   "IA Compressor Shutdown Active" : Bool = PLC "10 DI_DATA".E131_SHTDN AT %DB1.DBX0.0, 1 s
   "IDB_ATO2B_1_HIGH LEVEL VALUE (H)" : Real = PLC IDB_ATO2B_1."HIGH LEVEL VALUE (H)" AT %DB731.DBD30, 1 s
   "IDB_ATO2B_1_LOW LEVEL VALUE (L)" : Real = PLC IDB_ATO2B_1."LOW LEVEL VALUE (L)" AT %DB731.DBD26, 1 s
   "IDB_ATO2B_1_VERY HIGH LEVEL VALUE (HH)" : Real = PLC IDB_ATO2B_1."VERY HIGH LEVEL VALUE (HH)" AT %DB731.DBD34, 1 s
   "IDB_ATO2B_1_VERY LOW LEVEL VALUE (LL)" : Real = PLC IDB_ATO2B_1."VERY LOW LEVEL VALUE (LL)" AT %DB731.DBD22, 1 s
   "IDB_E-600_HIGH LEVEL VALUE (H)" : Real = PLC "IDB_E-600"."HIGH LEVEL VALUE (H)" AT %DB600.DBD30, 1 s
   "IDB_E-600_LOW LEVEL VALUE (L)" : Real = PLC "IDB_E-600"."LOW LEVEL VALUE (L)" AT %DB600.DBD26, 1 s
   "IDB_E-600_VERY HIGH LEVEL VALUE (HH)" : Real = PLC "IDB_E-600"."VERY HIGH LEVEL VALUE (HH)" AT %DB600.DBD34, 1 s
   "IDB_E-600_VERY LOW LEVEL VALUE (LL)" : Real = PLC "IDB_E-600"."VERY LOW LEVEL VALUE (LL)" AT %DB600.DBD22, 1 s
   "IDB_E700 Alarms_HIGH LEVEL VALUE (H)" : Real = PLC "IDB_E700 Alarms"."HIGH LEVEL VALUE (H)" AT %DB701.DBD30, 1 s
   "IDB_E700 Alarms_LOW LEVEL VALUE (L)" : Real = PLC "IDB_E700 Alarms"."LOW LEVEL VALUE (L)" AT %DB701.DBD26, 1 s
   "IDB_E700 Alarms_VERY HIGH LEVEL VALUE (HH)" : Real = PLC "IDB_E700 Alarms"."VERY HIGH LEVEL VALUE (HH)" AT %DB701.DBD34, 1 s
   "IDB_E700 Alarms_VERY LOW LEVEL VALUE (LL)" : Real = PLC "IDB_E700 Alarms"."VERY LOW LEVEL VALUE (LL)" AT %DB701.DBD22, 1 s
   "IDB_PIT 102_HIGH LEVEL VALUE (H)" : Real = PLC "IDB_PIT 102"."HIGH LEVEL VALUE (H)" AT %DB722.DBD30, 1 s
   "IDB_PIT 102_LOW LEVEL VALUE (L)" : Real = PLC "IDB_PIT 102"."LOW LEVEL VALUE (L)" AT %DB722.DBD26, 1 s
   "IDB_PIT 102_VERY HIGH LEVEL VALUE (HH)" : Real = PLC "IDB_PIT 102"."VERY HIGH LEVEL VALUE (HH)" AT %DB722.DBD34, 1 s
   "IDB_PIT 102_VERY LOW LEVEL VALUE (LL)" : Real = PLC "IDB_PIT 102"."VERY LOW LEVEL VALUE (LL)" AT %DB722.DBD22, 1 s
   "IDB_PIT 204_HIGH LEVEL VALUE (H)" : Real = PLC "IDB_PIT 204"."HIGH LEVEL VALUE (H)" AT %DB724.DBD30, 1 s
   "IDB_PIT 204_LOW LEVEL VALUE (L)" : Real = PLC "IDB_PIT 204"."LOW LEVEL VALUE (L)" AT %DB724.DBD26, 1 s
   "IDB_PIT 204_VERY HIGH LEVEL VALUE (HH)" : Real = PLC "IDB_PIT 204"."VERY HIGH LEVEL VALUE (HH)" AT %DB724.DBD34, 1 s
   "IDB_PIT 204_VERY LOW LEVEL VALUE (LL)" : Real = PLC "IDB_PIT 204"."VERY LOW LEVEL VALUE (LL)" AT %DB724.DBD22, 1 s
   "IDB_PIT 316_HIGH LEVEL VALUE (H)" : Real = PLC "IDB_PIT 316"."HIGH LEVEL VALUE (H)" AT %DB716.DBD30, 1 s
   "IDB_PIT 316_LOW LEVEL VALUE (L)" : Real = PLC "IDB_PIT 316"."LOW LEVEL VALUE (L)" AT %DB716.DBD26, 1 s
   "IDB_PIT 316_VERY HIGH LEVEL VALUE (HH)" : Real = PLC "IDB_PIT 316"."VERY HIGH LEVEL VALUE (HH)" AT %DB716.DBD34, 1 s
   "IDB_PIT 316_VERY LOW LEVEL VALUE (LL)" : Real = PLC "IDB_PIT 316"."VERY LOW LEVEL VALUE (LL)" AT %DB716.DBD22, 1 s
   "IDB_PIT 359_HIGH LEVEL VALUE (H)" : Real = PLC "IDB_PIT 359"."HIGH LEVEL VALUE (H)" AT %DB759.DBD30, 1 s
   "IDB_PIT 359_LOW LEVEL VALUE (L)" : Real = PLC "IDB_PIT 359"."LOW LEVEL VALUE (L)" AT %DB759.DBD26, 1 s
   "IDB_PIT 359_VERY HIGH LEVEL VALUE (HH)" : Real = PLC "IDB_PIT 359"."VERY HIGH LEVEL VALUE (HH)" AT %DB759.DBD34, 1 s
   "IDB_PIT 359_VERY LOW LEVEL VALUE (LL)" : Real = PLC "IDB_PIT 359"."VERY LOW LEVEL VALUE (LL)" AT %DB759.DBD22, 1 s
   "IDB_PIT 402_HIGH LEVEL VALUE (H)" : Real = PLC "IDB_PIT 402"."HIGH LEVEL VALUE (H)" AT %DB742.DBD30, 1 s
   "IDB_PIT 402_LOW LEVEL VALUE (L)" : Real = PLC "IDB_PIT 402"."LOW LEVEL VALUE (L)" AT %DB742.DBD26, 1 s
   "IDB_PIT 402_VERY HIGH LEVEL VALUE (HH)" : Real = PLC "IDB_PIT 402"."VERY HIGH LEVEL VALUE (HH)" AT %DB742.DBD34, 1 s
   "IDB_PIT 402_VERY LOW LEVEL VALUE (LL)" : Real = PLC "IDB_PIT 402"."VERY LOW LEVEL VALUE (LL)" AT %DB742.DBD22, 1 s
   "IDB_TIT 315_HIGH LEVEL VALUE (H)" : Real = PLC "IDB_TIT 315"."HIGH LEVEL VALUE (H)" AT %DB715.DBD30, 1 s
   "IDB_TIT 315_LOW LEVEL VALUE (L)" : Real = PLC "IDB_TIT 315"."LOW LEVEL VALUE (L)" AT %DB715.DBD26, 1 s
   "IDB_TIT 315_VERY HIGH LEVEL VALUE (HH)" : Real = PLC "IDB_TIT 315"."VERY HIGH LEVEL VALUE (HH)" AT %DB715.DBD34, 1 s
   "IDB_TIT 315_VERY LOW LEVEL VALUE (LL)" : Real = PLC "IDB_TIT 315"."VERY LOW LEVEL VALUE (LL)" AT %DB715.DBD22, 1 s
   "IDB_TIT 319_HIGH LEVEL VALUE (H)" : Real = PLC "IDB_TIT 319"."HIGH LEVEL VALUE (H)" AT %DB719.DBD30, 1 s
   "IDB_TIT 319_LOW LEVEL VALUE (L)" : Real = PLC "IDB_TIT 319"."LOW LEVEL VALUE (L)" AT %DB719.DBD26, 1 s
   "IDB_TIT 319_VERY HIGH LEVEL VALUE (HH)" : Real = PLC "IDB_TIT 319"."VERY HIGH LEVEL VALUE (HH)" AT %DB719.DBD34, 1 s
   "IDB_TIT 319_VERY LOW LEVEL VALUE (LL)" : Real = PLC "IDB_TIT 319"."VERY LOW LEVEL VALUE (LL)" AT %DB719.DBD22, 1 s
   "IDB_TIT 360_HIGH LEVEL VALUE (H)" : Real = PLC "IDB_TIT 360"."HIGH LEVEL VALUE (H)" AT %DB760.DBD30, 1 s
   "IDB_TIT 360_LOW LEVEL VALUE (L)" : Real = PLC "IDB_TIT 360"."LOW LEVEL VALUE (L)" AT %DB760.DBD26, 1 s
   "IDB_TIT 360_VERY HIGH LEVEL VALUE (HH)" : Real = PLC "IDB_TIT 360"."VERY HIGH LEVEL VALUE (HH)" AT %DB760.DBD34, 1 s
   "IDB_TIT 360_VERY LOW LEVEL VALUE (LL)" : Real = PLC "IDB_TIT 360"."VERY LOW LEVEL VALUE (LL)" AT %DB760.DBD22, 1 s
   "IDB_TIT 401_HIGH LEVEL VALUE (H)" : Real = PLC "IDB_TIT 401"."HIGH LEVEL VALUE (H)" AT %DB741.DBD30, 1 s
   "IDB_TIT 401_LOW LEVEL VALUE (L)" : Real = PLC "IDB_TIT 401"."LOW LEVEL VALUE (L)" AT %DB741.DBD26, 1 s
   "IDB_TIT 401_VERY HIGH LEVEL VALUE (HH)" : Real = PLC "IDB_TIT 401"."VERY HIGH LEVEL VALUE (HH)" AT %DB741.DBD34, 1 s
   "IDB_TIT 401_VERY LOW LEVEL VALUE (LL)" : Real = PLC "IDB_TIT 401"."VERY LOW LEVEL VALUE (LL)" AT %DB741.DBD22, 1 s
   "IG Press SP (R)" : Real = PLC "19_AUTO_CMNDS_Data".PIT402_Target AT %DB1.DBD0, 1 s
   "IG Shell Temp Hi Switch" : Bool = PLC "10 DI_DATA".TS006 AT %DB1.DBX0.0, 1 s
   "IG Soot Content Scaled" : Real = PLC "12_AI_Data".E700SootContentIn AT %DB1.DBX0.0, 1 s
   "IG Temp Hi Hi Switch" : Bool = PLC "10 DI_DATA".TS403_FAULT AT %DB1.DBX0.0, 1 s
   "IG Temperature High (TS403)" : Bool = PLC "10 DI_DATA".TS403_FAULT AT %DB1.DBX0.0, 1 s
   "IGG Automated" : Bool = PLC "80_From_HMI".Request_Auto AT %DB1.DBX0.0, 1 s
   "IGG E-Stop Healthy" : Bool = PLC "10_DI_Data".IGG_ESTOP_OK AT %DB1.DBX0.0, 1 s
   "IGG Inlet Fuel Pressure (PIT204) Scaled" : Real = PLC "12_AI_Data".PIT204In_SCALED AT %DB1.DBX0.0, 1 s
   "IGG Inlet Fuel Temp (TIT202) Scaled" : Real = PLC "12_AI_Data".TIT202In_SCALED AT %DB1.DBX0.0, 1 s
   "IGG Main Atom Air Presure (PIT113) Scaled" : Real = PLC "12_AI_Data".PIT113In_SCALED AT %DB1.DBX0.0, 1 s
   "IGG Main Fuel Pressure (PIT205) Scaled" : Real = PLC "12_AI_Data".PIT205In_SCALED AT %DB1.DBX0.0, 1 s
   "IGG Manual" : Bool = PLC "80_From_HMI".Request_Manual AT %DB1.DBX0.0, 1 s
   "IGG Running" : Bool = PLC "14_DQ_Data".24PF1 AT %DB1.DBX0.0, 1 s
   "IGG Shell High Temp (TS006)" : Bool = PLC "10 DI_DATA".TS006 AT %DB1.DBX0.0, 1 s
   "IGG Shutdown Alarm Active" : Bool = PLC "14_DQ_Data".24K3 AT %DB1.DBX0.0, 1 s
   "IGG Shutting Down animation" : Bool = PLC "14_DQ_Data".24K3 AT %DB1.DBX0.0, 1 s
   "IGG Start Warning" : Bool = PLC "Sequence Times_DB"."Warn to IGG Start" AT %DB1.DBW0, 1 s
   "IGG Vent Power Healthy" : Bool = PLC "10_DI_Data".IGG_VNT_PWR_OK AT %DB1.DBX0.0, 1 s
   "IGG Warning Alarm Active" : Bool = PLC "14_DQ_Data".24K4 AT %DB1.DBX0.0, 1 s
   "IGG_Step_Time_001" : Time = PLC "86_Times".STEP_MAX_TIME_STP_001 AT %DB1.DBW0, 1 s
   "IGG_Step_Time_005" : Time = PLC "86_Times".STEP_MAX_TIME_STP_005 AT %DB1.DBW0, 1 s
   "IGG_Step_Time_010" : Time = PLC "86_Times".STEP_MAX_TIME_STP_010 AT %DB1.DBW0, 1 s
   "IGG_Step_Time_020" : Time = PLC "86_Times".STEP_MAX_TIME_STP_020 AT %DB1.DBW0, 1 s
   "IGG_Step_Time_030" : Time = PLC "86_Times".STEP_MAX_TIME_STP_030 AT %DB1.DBW0, 1 s
   "IGG_Step_Time_040" : Time = PLC "86_Times".STEP_MAX_TIME_STP_040 AT %DB1.DBW0, 1 s
   "IGG_Step_Time_050" : Time = PLC "86_Times".STEP_MAX_TIME_STP_050 AT %DB1.DBW0, 1 s
   "IGG_Step_Time_060" : Time = PLC "86_Times".STEP_MAX_TIME_STP_060 AT %DB1.DBW0, 1 s
   "IGG_Step_Time_070" : Time = PLC "86_Times".STEP_MAX_TIME_STP_070 AT %DB1.DBW0, 1 s
   "IGG_Step_Time_080" : Time = PLC "86_Times".STEP_MAX_TIME_STP_080 AT %DB1.DBW0, 1 s
   "IGG_Step_Time_090" : Time = PLC "86_Times".STEP_MAX_TIME_STP_090 AT %DB1.DBW0, 1 s
   "IGG_Step_Time_100" : Time = PLC "86_Times".STEP_MAX_TIME_STP_100 AT %DB1.DBW0, 1 s
   "IGG_Step_Time_110" : Time = PLC "86_Times".STEP_MAX_TIME_STP_110 AT %DB1.DBW0, 1 s
   "IGG_Step_Time_120" : Time = PLC "86_Times".STEP_MAX_TIME_STP_120 AT %DB1.DBW0, 1 s
   "IGG_Step_Time_130" : Time = PLC "86_Times".STEP_MAX_TIME_STP_130 AT %DB1.DBW0, 1 s
   "IGG_Step_Time_140" : Time = PLC "86_Times".STEP_MAX_TIME_STP_140 AT %DB1.DBW0, 1 s
   "IGG_Step_Time_150" : Time = PLC "86_Times".STEP_MAX_TIME_STP_150 AT %DB1.DBW0, 1 s
   "IGG_Step_Time_160" : Time = PLC "86_Times".STEP_MAX_TIME_STP_160 AT %DB1.DBW0, 1 s
   "IGG_Step_Time_170" : Time = PLC "86_Times".STEP_MAX_TIME_STP_170 AT %DB1.DBW0, 1 s
   "IGG_Step_Time_180" : Time = PLC "86_Times".STEP_MAX_TIME_STP_180 AT %DB1.DBW0, 1 s
   "IGG_Step_Time_190" : Time = PLC "86_Times".STEP_MAX_TIME_STP_190 AT %DB1.DBW0, 1 s
   "IGG_Step_Time_200" : Time = PLC "86_Times".STEP_MAX_TIME_STP_200 AT %DB1.DBW0, 1 s
   "IGG_Step_Time_210" : Time = PLC "86_Times".STEP_MAX_TIME_STP_210 AT %DB1.DBW0, 1 s
   "IGG_Step_Time_220" : Time = PLC "86_Times".STEP_MAX_TIME_STP_220 AT %DB1.DBW0, 1 s
   "IGG_Step_Time_230" : Time = PLC "86_Times".STEP_MAX_TIME_STP_230 AT %DB1.DBW0, 1 s
   "IGG_Step_Time_240" : Time = PLC "86_Times".STEP_MAX_TIME_STP_240 AT %DB1.DBW0, 1 s
   "IGG_Step_Time_250" : Time = PLC "86_Times".STEP_MAX_TIME_STP_250 AT %DB1.DBW0, 1 s
   "IGG_Step_Time_260" : Time = PLC "86_Times".STEP_MAX_TIME_STP_260 AT %DB1.DBW0, 1 s
   "IGG_Step_Time_270" : Time = PLC "86_Times".STEP_MAX_TIME_STP_270 AT %DB1.DBW0, 1 s
   "IGG_Step_Time_280" : Time = PLC "86_Times".STEP_MAX_TIME_STP_280 AT %DB1.DBW0, 1 s
   "IGG_Step_Time_290" : Time = PLC "86_Times".STEP_MAX_TIME_STP_290 AT %DB1.DBW0, 1 s
   "IGG_Step_Time_300" : Time = PLC "86_Times".STEP_MAX_TIME_STP_300 AT %DB1.DBW0, 1 s
   "IGG_Step_Time_310" : Time = PLC "86_Times".STEP_MAX_TIME_STP_310 AT %DB1.DBW0, 1 s
   "IGG_Step_Time_320" : Time = PLC "86_Times".STEP_MAX_TIME_STP_320 AT %DB1.DBW0, 1 s
   "IGG_Step_Time_330" : Time = PLC "86_Times".STEP_MAX_TIME_STP_330 AT %DB1.DBW0, 1 s
   "IGG_Step_Time_340" : Time = PLC "86_Times".STEP_MAX_TIME_STP_340 AT %DB1.DBW0, 1 s
   "IGG_Step_Time_350" : Time = PLC "86_Times".STEP_MAX_TIME_STP_350 AT %DB1.DBW0, 1 s
   "IGG_Step_Time_360" : Time = PLC "86_Times".STEP_MAX_TIME_STP_360 AT %DB1.DBW0, 1 s
   "IGG_Step_Time_370" : Time = PLC "86_Times".STEP_MAX_TIME_STP_370 AT %DB1.DBW0, 1 s
   "IGG_Step_Time_380" : Time = PLC "86_Times".STEP_MAX_TIME_STP_380 AT %DB1.DBW0, 1 s
   "IGG_Step_Time_390" : Time = PLC "86_Times".STEP_MAX_TIME_STP_390 AT %DB1.DBW0, 1 s
   "IGG_Step_Time_400" : Time = PLC "86_Times".STEP_MAX_TIME_STP_400 AT %DB1.DBW0, 1 s
   "IGG_Step_Time_410" : Time = PLC "86_Times".STEP_MAX_TIME_STP_410 AT %DB1.DBW0, 1 s
   "IGG_Step_Time_420" : Time = PLC "86_Times".STEP_MAX_TIME_STP_420 AT %DB1.DBW0, 1 s
   "IGG_Step_Time_430" : Time = PLC "86_Times".STEP_MAX_TIME_STP_430 AT %DB1.DBW0, 1 s
   "IGG_Step_Time_440" : Time = PLC "86_Times".STEP_MAX_TIME_STP_440 AT %DB1.DBW0, 1 s
   "IGG_Step_Time_450" : Time = PLC "86_Times".STEP_MAX_TIME_STP_450 AT %DB1.DBW0, 1 s
   "IGG_Step_Time_460" : Time = PLC "86_Times".STEP_MAX_TIME_STP_460 AT %DB1.DBW0, 1 s
   "IGG_Step_Time_470" : Time = PLC "86_Times".STEP_MAX_TIME_STP_470 AT %DB1.DBW0, 1 s
   "IGG_Step_Time_480" : Time = PLC "86_Times".STEP_MAX_TIME_STP_480 AT %DB1.DBW0, 1 s
   "IGG_Step_Time_490" : Time = PLC "86_Times".STEP_MAX_TIME_STP_490 AT %DB1.DBW0, 1 s
   "IGG_Step_Time_500" : Time = PLC "86_Times".STEP_MAX_TIME_STP_500 AT %DB1.DBW0, 1 s
   "IGG_Times_Burner Control Start Command Delay" : Time = PLC "86_Times".PRE_BC_STRT_CMND_DLY AT %DB1.DBD0, 1 s
   "IGG_Times_CV203 Close Command" : Time = PLC "86_Times".PRE_CV203_CLS_CMND_DLY AT %DB1.DBD0, 1 s
   "IGG_Times_CV311 Max" : Time = PLC "86_Times".CV311_MAX_TRVL_TIME AT %DB1.DBD0, 1 s
   "IGG_Times_CV312 Max" : Time = PLC "86_Times".CV312_MAX_TRVL_TIME AT %DB1.DBD0, 1 s
   "IGG_Times_CV321 Max" : Time = PLC "86_Times".CV321_MAX_TRVL_TIME AT %DB1.DBD0, 1 s
   "IGG_Times_CV322 Max" : Time = PLC "86_Times".CV322_MAX_TRVL_TIME AT %DB1.DBD0, 1 s
   "IGG_Times_CV401 Max" : Time = PLC "86_Times".CV401_MAX_TRVL_TIME AT %DB1.DBD0, 1 s
   "IGG_Times_CV431 Max" : Time = PLC "86_Times".CV431_MAX_TRVL_TIME AT %DB1.DBD0, 1 s
   "IGG_Times_CV432 Max" : Time = PLC "86_Times".CV432_MAX_TRVL_TIME AT %DB1.DBD0, 1 s
   "IGG_Times_Post CV311 Close" : Time = PLC "86_Times".POST_CV311_CLS_DLY AT %DB1.DBD0, 1 s
   "IGG_Times_Post CV321 Open" : Time = PLC "86_Times".POST_CV321_OPN_DLY AT %DB1.DBD0, 1 s
   "IGG_Times_Post P301 Stop" : Time = PLC "86_Times".POST_P301_STOP_DLY AT %DB1.DBD0, 1 s
   "Igniter Control" : Bool = PLC "14_DQ_Data".X001ControlOut AT %DB1.DBX0.0, 1 s
   "Ignitor Power Healthy" : Bool = PLC "10 DI_DATA".X001_PWR_OK AT %DB1.DBX0.0, 1 s
   "Inert Gas Pressure (PIT402) Scaled" : Real = PLC "12_AI_Data".PIT402_SCALED AT %DB1.DBX0.0, 1 s
   "Inert Gas Temp Scaled" : Real = PLC "12_AI_Data".TIT401_SCALED AT %DB1.DBX0.0, 1 s
   "Inlet CSW Pressured PIT359 Scaled" : Real = PLC "12_AI_Data".PIT359_SCALED AT %DB1.DBX0.0, 1 s
   "Inlet CSW Temp Scaled" : Real = PLC "12_AI_Data".TIT319_SCALED AT %DB1.DBX0.0, 1 s
   "Inlet IA Pressure PIT112 Scaled" : Real = PLC "12_AI_Data".PIT112In_SCALED AT %DB1.DBX0.0, 1 s
   "Jacket Cooling Water Flow Switch" : Bool = PLC "10 DI_DATA".FS317 AT %DB1.DBX0.0, 1 s
   "LIT304_ALM_ANALOG_DB71_HIGH LEVEL VALUE (H)" : Real = PLC LIT304_ALM_ANALOG_DB71."HIGH LEVEL VALUE (H)" AT %DB71.DBD30, 1 s
   "LIT304_ALM_ANALOG_DB71_LOW LEVEL VALUE (L)" : Real = PLC LIT304_ALM_ANALOG_DB71."LOW LEVEL VALUE (L)" AT %DB71.DBD26, 1 s
   "LIT304_ALM_ANALOG_DB71_VERY HIGH LEVEL VALUE (HH)" : Real = PLC LIT304_ALM_ANALOG_DB71."VERY HIGH LEVEL VALUE (HH)" AT %DB71.DBD34, 1 s
   "LIT304_ALM_ANALOG_DB71_VERY LOW LEVEL VALUE (LL)" : Real = PLC LIT304_ALM_ANALOG_DB71."VERY LOW LEVEL VALUE (LL)" AT %DB71.DBD22, 1 s
   "Logging SD Card Overflow" : Bool AT %DB1.DBX0.0
      on ChangeValue: "SD_Card_Overflow"()
   "Main Atom Air Flow  OK" : Bool = PLC "10 DI_DATA".FS115 AT %DB1.DBX0.0, 1 s
   "Main Atom Air Flow Switch" : Bool = PLC "10 DI_DATA".FS115 AT %DB1.DBW0, 1 s
   "Main Atom Air Reg Valve Position" : Real = PLC "16_AQ_Data".CV111_CNTRL AT %DB1.DBD0, 1 s
   "Main B Atom Air Valve Control" : Bool = PLC "14_DQ_Data".200CV114ControlOut AT %DB1.DBX0.0, 1 s
   "Main B Fuel Valve 1 Control" : Bool = PLC "14_DQ_Data".200CV206ControlOut AT %DB1.DBX0.0, 1 s
   "Main B Fuel Valve 2 Control" : Bool = PLC "14_DQ_Data".200CV207ControlOut AT %DB1.DBX0.0, 1 s
   "Main Fuel Reg Valve Control" : Real = PLC "16_AQ_Data".CV203_CNTRL AT %DB1.DBD0, 1 s
   "Main Fuel Reg Valve Position" : Real = PLC "16_AQ_Data".CV203_CNTRL, 1 s
   "Maintained 24V Power" : Bool = PLC "10_DI_Data".MAINTD_24VDC_PWR_OK AT %DB1.DBX0.0, 1 s
   "MAN_AQ100_DEC_CAB_Speed" : Bool = PLC "80_From_HMI".MAN_AQ_DEC_100 AT %DB1.DBX0.0, 1 s
   "MAN_AQ100_DEC_Main_Fuel_Reg" : Bool = PLC "80_From_HMI".MAN_AQ_DEC_100 AT %DB1.DBX0.0, 1 s
   "MAN_AQ100_INC_CAB_Speed" : Bool = PLC "80_From_HMI".MAN_AQ_INC_100 AT %DB1.DBX0.0, 1 s
   "MAN_AQ100_INC_Main_Fuel_Reg" : Bool = PLC "80_From_HMI".MAN_AQ_INC_100 AT %DB1.DBX0.0, 1 s
   "MAN_AQ102_DEC_Main_Atom_Air" : Bool = PLC "80_From_HMI".MAN_AQ_DEC_102 AT %DB1.DBX0.0, 1 s
   "MAN_AQ102_DEC_SPARE" : Bool = PLC "80_From_HMI".MAN_AQ_DEC_102 AT %DB1.DBX0.0, 1 s
   "MAN_AQ102_INC_Main_Atom_Air" : Bool = PLC "80_From_HMI".MAN_AQ_INC_102 AT %DB1.DBX0.0, 1 s
   "MAN_AQ102_INC_SPARE" : Bool = PLC "80_From_HMI".MAN_AQ_INC_102 AT %DB1.DBX0.0, 1 s
   "MAN_AQ104_DEC_SPARE" : Bool = PLC "80_From_HMI".MAN_AQ_DEC_104 AT %DB1.DBX0.0, 1 s
   "MAN_AQ104_INC_SPARE" : Bool = PLC "80_From_HMI".MAN_AQ_INC_104 AT %DB1.DBX0.0, 1 s
   "MAN_AQ96_DEC_SPARE" : Bool = PLC "80_From_HMI".MAN_AQ_DEC_96 AT %DB1.DBX0.0, 1 s
   "MAN_AQ96_INC_SPARE" : Bool = PLC "80_From_HMI".MAN_AQ_INC_96 AT %DB1.DBX0.0, 1 s
   "MAN_AQ98_DEC_SPARE" : Bool = PLC "80_From_HMI".MAN_AQ_DEC_98 AT %DB1.DBX0.0, 1 s
   "MAN_AQ98_DEC_Vent_Valve_Pos" : Bool = PLC "80_From_HMI".MAN_AQ_DEC_98 AT %DB1.DBX0.0, 1 s
   "MAN_AQ98_INC_SPARE" : Bool = PLC "80_From_HMI".MAN_AQ_INC_98 AT %DB1.DBX0.0, 1 s
   "MAN_AQ98_INC_Vent_Valve_Pos" : Bool = PLC "80_From_HMI".MAN_AQ_INC_98 AT %DB1.DBX0.0, 1 s
   "MAN_Q0.0_FP1" : Bool = PLC "80_From_HMI".MAN_DQ_0_0 AT %DB1.DBX0.0, 1 s
   "MAN_Q0.0_Test_Press" : Bool = PLC "80_From_HMI".MAN_DQ_0_0 AT %DB1.DBX0.0, 1 s
   "MAN_Q0.1_FP2" : Bool = PLC "80_From_HMI".MAN_DQ_0_1 AT %DB1.DBX0.0, 1 s
   "MAN_Q0.1_Pilot_IGN" : Bool = PLC "80_From_HMI".MAN_DQ_0_1 AT %DB1.DBX0.0, 1 s
   "MAN_Q0.2_CAB" : Bool = PLC "80_From_HMI".MAN_DQ_0_2 AT %DB1.DBX0.0, 1 s
   "MAN_Q0.2_PilotFuel1" : Bool = PLC "80_From_HMI".MAN_DQ_0_2 AT %DB1.DBX0.0, 1 s
   "MAN_Q0.3_CSW_Inlet" : Bool = PLC "80_From_HMI".MAN_DQ_0_3 AT %DB1.DBX0.0, 1 s
   "MAN_Q0.3_PilotFuel2" : Bool = PLC "80_From_HMI".MAN_DQ_0_3 AT %DB1.DBX0.0, 1 s
   "MAN_Q0.4_CSW_Drain" : Bool = PLC "80_From_HMI".MAN_DQ_0_4 AT %DB1.DBX0.0, 1 s
   "MAN_Q0.4_MainAtom" : Bool = PLC "80_From_HMI".MAN_DQ_0_4 AT %DB1.DBX0.0, 1 s
   "MAN_Q0.5_IGSupply" : Bool = PLC "80_From_HMI".MAN_DQ_0_5 AT %DB1.DBX0.0, 1 s
   "MAN_Q0.5_MainFuel1" : Bool = PLC "80_From_HMI".MAN_DQ_0_5 AT %DB1.DBX0.0, 1 s
   "MAN_Q0.6_CB/BWTS" : Bool = PLC "80_From_HMI".MAN_DQ_0_6 AT %DB1.DBX0.0, 1 s
   "MAN_Q0.6_MainFuel2" : Bool = PLC "80_From_HMI".MAN_DQ_0_6 AT %DB1.DBX0.0, 1 s
   "MAN_Q0.7_IAComp" : Bool = PLC "80_From_HMI".MAN_DQ_0_7 AT %DB1.DBX0.0, 1 s
   "MAN_Q0.7_Spare" : Bool = PLC "80_From_HMI".MAN_DQ_0_7 AT %DB1.DBX0.0, 1 s
   "MAN_Q1.0_CSWPump" : Bool = PLC "80_From_HMI".MAN_DQ_1_0 AT %DB1.DBX0.0, 1 s
   "MAN_Q1.0_Spare" : Bool = PLC "80_From_HMI".MAN_DQ_1_0 AT %DB1.DBX0.0, 1 s
   "MAN_Q1.1_Atmos" : Bool = PLC "80_From_HMI".MAN_DQ_1_1 AT %DB1.DBX0.0, 1 s
   "MAN_Q1.1_IGN" : Bool = PLC "80_From_HMI".MAN_DQ_1_1 AT %DB1.DBX0.0, 1 s
   "MAN_Q1.2_IGG_SD" : Bool = PLC "80_From_HMI".MAN_DQ_1_2 AT %DB1.DBX0.0, 1 s
   "MAN_Q1.2_Spare" : Bool = PLC "80_From_HMI".MAN_DQ_1_2 AT %DB1.DBX0.0, 1 s
   "MAN_Q1.3_IGG_WRN" : Bool = PLC "80_From_HMI".MAN_DQ_1_3 AT %DB1.DBX0.0, 1 s
   "MAN_Q1.3_Spare" : Bool = PLC "80_From_HMI".MAN_DQ_1_3 AT %DB1.DBX0.0, 1 s
   "MAN_Q1.4_IGG_RNG" : Bool = PLC "80_From_HMI".MAN_DQ_1_4 AT %DB1.DBX0.0, 1 s
   "MAN_Q1.4_Spare" : Bool = PLC "80_From_HMI".MAN_DQ_1_4 AT %DB1.DBX0.0, 1 s
   "MAN_Q1.5_SD" : Bool = PLC "80_From_HMI".MAN_DQ_1_5 AT %DB1.DBX0.0, 1 s
   "MAN_Q1.5_Spare" : Bool = PLC "80_From_HMI".MAN_DQ_1_5 AT %DB1.DBX0.0, 1 s
   "MAN_Q1.6_Spare" : Bool = PLC "80_From_HMI".MAN_DQ_1_6 AT %DB1.DBX0.0, 1 s
   "MAN_Q1.6_WRN" : Bool = PLC "80_From_HMI".MAN_DQ_1_6 AT %DB1.DBX0.0, 1 s
   "MAN_Q1.7_BUZ" : Bool = PLC "80_From_HMI".MAN_DQ_1_7 AT %DB1.DBX0.0, 1 s
   "MAN_Q1.7_CSW_Pump" : Bool = PLC "80_From_HMI".MAN_DQ_1_7 AT %DB1.DBX0.0, 1 s
   "MCC Vent Power Healthy" : Bool = PLC "10_DI_Data".MCC_VNT_PWR_OK AT %DB1.DBX0.0, 1 s
   "Not BWT mode Warning" : Bool = PLC "2068_Sys_Status_Data"."Not BWT mode Warning" AT %DB1.DBD0, 1 s
   "Nozzle Cooling Water Flow Switch" : Bool = PLC "10 DI_DATA".FS320 AT %DB1.DBX0.0, 1 s
   "O2 Analyser Content Scaled" : Real = PLC "12_AI_Data".E600O2ContentIn AT %DB1.DBX0.0, 100 ms
   "O2 Analyser Hi Hi" : Bool = PLC "10 DI_DATA".E600_HIHI AT %DB1.DBX0.0, 1 s
   "O2 Analyser Lo Lo" : Bool = PLC "10 DI_DATA".E600_LOLO AT %DB1.DBX0.0, 1 s
   "O2 Ramp Control_QLMN_HLM" : Bool = PLC "O2 Ramp Control".QLMN_HLM, 1 s
   "O2 Ramp Control_QLMN_LLM" : Bool = PLC "O2 Ramp Control".QLMN_LLM, 1 s
   "O2 System Fail" : Bool = PLC "10 DI_DATA".E600_NOK AT %DB1.DBX0.0, 1 s
   "O2 System Power Healthy" : Bool = PLC "10 DI_DATA".E600_PWR_OK AT %DB1.DBX0.0, 1 s
   "Operation hours E139_IDB_Hours Functioning" : Int = PLC "Operation hours E139_IDB"."Hours Functioning", 1 s
   "Outlet CSW Pressure PIT316 Scaled" : Real = PLC "12_AI_Data".PIT316_SCALED AT %DB1.DBX0.0, 1 s
   "Outlet CSW Temp Scaled" : Real = PLC "12_AI_Data".TIT360_SCALED AT %DB1.DBX0.0, 1 s
   "P301 Present" : Bool = PLC "80_From_HMI".P301_PRSNT AT %DB1.DBX0.0, 1 s
   "P305_Functioning Hours_IDB_Hours Functioning Out" : Int = PLC "P305_Functioning Hours_IDB"."Hours Functioning Out", 1 s
   "PGC_COMMISSION_MODE_DB_Active" : Bool = PLC PGC_COMMISSION_MODE_DB.Active, 1 s
   "PGC_COMMISSION_MODE_DB_Button Control" : Int = PLC PGC_COMMISSION_MODE_DB."Button Control", 1 s
   "PGC_COMMISSION_MODE_DB_Drive Popup" : Bool = PLC PGC_COMMISSION_MODE_DB."Drive Popup", 500 ms
   "PGC_COMMISSION_MODE_DB_Setpoint" : Real = PLC PGC_COMMISSION_MODE_DB.Setpoint, 1 s
   "Pilot Air Flow  OK" : Bool = PLC "10 DI_DATA".FS123 AT %DB1.DBX0.0, 1 s
   "Pilot B Fuel Valve 1 Control" : Bool = PLC "14_DQ_Data".200CV215ControlOut AT %DB1.DBX0.0, 1 s
   "Pilot B Fuel Valve 2 Control" : Bool = PLC "14_DQ_Data".200CV216ControlOut AT %DB1.DBX0.0, 1 s
   "Pilot B Ignition Air Valve Control" : Bool = PLC "14_DQ_Data".200CV124ControlOut AT %DB1.DBX0.0, 1 s
   "Pilot Flame" : Bool = PLC "102_Pilot_Burner_DB".FLM_DET AT %DB1.DBX0.0, 100 ms
   "PilotPurgeOK" : Bool = PLC "104_Pilot_Purge_DB".DN_OK AT %DB1.DBX0.0, 1 s
   "PIT348_ALM_ANALOG_DB73_HIGH LEVEL VALUE (H)" : Real = PLC PIT348_ALM_ANALOG_DB73."HIGH LEVEL VALUE (H)" AT %DB73.DBD30, 1 s
   "PIT348_ALM_ANALOG_DB73_LOW LEVEL VALUE (L)" : Real = PLC PIT348_ALM_ANALOG_DB73."LOW LEVEL VALUE (L)" AT %DB73.DBD26, 1 s
   "PIT348_ALM_ANALOG_DB73_VERY HIGH LEVEL VALUE (HH)" : Real = PLC PIT348_ALM_ANALOG_DB73."VERY HIGH LEVEL VALUE (HH)" AT %DB73.DBD34, 1 s
   "PIT348_ALM_ANALOG_DB73_VERY LOW LEVEL VALUE (LL)" : Real = PLC PIT348_ALM_ANALOG_DB73."VERY LOW LEVEL VALUE (LL)" AT %DB73.DBD22, 1 s
   "PIT353_ALM_ANALOG_DB72_HIGH LEVEL VALUE (H)" : Real = PLC PIT353_ALM_ANALOG_DB72."HIGH LEVEL VALUE (H)" AT %DB72.DBD30, 1 s
   "PIT353_ALM_ANALOG_DB72_LOW LEVEL VALUE (L)" : Real = PLC PIT353_ALM_ANALOG_DB72."LOW LEVEL VALUE (L)" AT %DB72.DBD26, 1 s
   "PIT353_ALM_ANALOG_DB72_VERY HIGH LEVEL VALUE (HH)" : Real = PLC PIT353_ALM_ANALOG_DB72."VERY HIGH LEVEL VALUE (HH)" AT %DB72.DBD34, 1 s
   "PIT353_ALM_ANALOG_DB72_VERY LOW LEVEL VALUE (LL)" : Real = PLC PIT353_ALM_ANALOG_DB72."VERY LOW LEVEL VALUE (LL)" AT %DB72.DBD22, 1 s
   "PIT358_ALM_ANALOG_DB78_HIGH LEVEL VALUE (H)" : Real = PLC PIT358_ALM_ANALOG_DB78."HIGH LEVEL VALUE (H)" AT %DB78.DBD30, 1 s
   "PIT358_ALM_ANALOG_DB78_LOW LEVEL VALUE (L)" : Real = PLC PIT358_ALM_ANALOG_DB78."LOW LEVEL VALUE (L)" AT %DB78.DBD26, 1 s
   "PIT358_ALM_ANALOG_DB78_VERY HIGH LEVEL VALUE (HH)" : Real = PLC PIT358_ALM_ANALOG_DB78."VERY HIGH LEVEL VALUE (HH)" AT %DB78.DBD34, 1 s
   "PIT358_ALM_ANALOG_DB78_VERY LOW LEVEL VALUE (LL)" : Real = PLC PIT358_ALM_ANALOG_DB78."VERY LOW LEVEL VALUE (LL)" AT %DB78.DBD22, 1 s
   "PIT424_RIO1_ALM_ANALOG_DB_HIGH LEVEL VALUE (H)" : Real = PLC PIT424_RIO1_ALM_ANALOG_DB."HIGH LEVEL VALUE (H)" AT %DB2219.DBD30, 1 s
   "PIT424_RIO1_ALM_ANALOG_DB_LOW LEVEL VALUE (L)" : Real = PLC PIT424_RIO1_ALM_ANALOG_DB."LOW LEVEL VALUE (L)" AT %DB2219.DBD26, 1 s
   "PIT424_RIO1_ALM_ANALOG_DB_VERY HIGH LEVEL VALUE (HH)" : Real = PLC PIT424_RIO1_ALM_ANALOG_DB."VERY HIGH LEVEL VALUE (HH)" AT %DB2219.DBD34, 1 s
   "PIT424_RIO1_ALM_ANALOG_DB_VERY LOW LEVEL VALUE (LL)" : Real = PLC PIT424_RIO1_ALM_ANALOG_DB."VERY LOW LEVEL VALUE (LL)" AT %DB2219.DBD22, 1 s
   "PIT424_RIO3_ALM_ANALOG_DB_HIGH LEVEL VALUE (H)" : Real = PLC PIT424_RIO3_ALM_ANALOG_DB."HIGH LEVEL VALUE (H)" AT %DB2220.DBD30, 1 s
   "PIT424_RIO3_ALM_ANALOG_DB_LOW LEVEL VALUE (L)" : Real = PLC PIT424_RIO3_ALM_ANALOG_DB."LOW LEVEL VALUE (L)" AT %DB2220.DBD26, 1 s
   "PIT424_RIO3_ALM_ANALOG_DB_VERY HIGH LEVEL VALUE (HH)" : Real = PLC PIT424_RIO3_ALM_ANALOG_DB."VERY HIGH LEVEL VALUE (HH)" AT %DB2220.DBD34, 1 s
   "PIT424_RIO3_ALM_ANALOG_DB_VERY LOW LEVEL VALUE (LL)" : Real = PLC PIT424_RIO3_ALM_ANALOG_DB."VERY LOW LEVEL VALUE (LL)" AT %DB2220.DBD22, 1 s
   "PIT424_RIO4_ALM_ANALOG_DB_HIGH LEVEL VALUE (H)" : Real = PLC PIT424_RIO4_ALM_ANALOG_DB."HIGH LEVEL VALUE (H)" AT %DB2221.DBD30, 1 s
   "PIT424_RIO4_ALM_ANALOG_DB_LOW LEVEL VALUE (L)" : Real = PLC PIT424_RIO4_ALM_ANALOG_DB."LOW LEVEL VALUE (L)" AT %DB2221.DBD26, 1 s
   "PIT424_RIO4_ALM_ANALOG_DB_VERY HIGH LEVEL VALUE (HH)" : Real = PLC PIT424_RIO4_ALM_ANALOG_DB."VERY HIGH LEVEL VALUE (HH)" AT %DB2221.DBD34, 1 s
   "PIT424_RIO4_ALM_ANALOG_DB_VERY LOW LEVEL VALUE (LL)" : Real = PLC PIT424_RIO4_ALM_ANALOG_DB."VERY LOW LEVEL VALUE (LL)" AT %DB2221.DBD22, 1 s
   "PIT424_RIO5_ALM_ANALOG_DB_HIGH LEVEL VALUE (H)" : Real = PLC PIT424_RIO5_ALM_ANALOG_DB."HIGH LEVEL VALUE (H)" AT %DB2222.DBD30, 1 s
   "PIT424_RIO5_ALM_ANALOG_DB_LOW LEVEL VALUE (L)" : Real = PLC PIT424_RIO5_ALM_ANALOG_DB."LOW LEVEL VALUE (L)" AT %DB2222.DBD26, 1 s
   "PIT424_RIO5_ALM_ANALOG_DB_VERY HIGH LEVEL VALUE (HH)" : Real = PLC PIT424_RIO5_ALM_ANALOG_DB."VERY HIGH LEVEL VALUE (HH)" AT %DB2222.DBD34, 1 s
   "PIT424_RIO5_ALM_ANALOG_DB_VERY LOW LEVEL VALUE (LL)" : Real = PLC PIT424_RIO5_ALM_ANALOG_DB."VERY LOW LEVEL VALUE (LL)" AT %DB2222.DBD22, 1 s
   "PIT424_RIO6_ALM_ANALOG_DB_HIGH LEVEL VALUE (H)" : Real = PLC PIT424_RIO6_ALM_ANALOG_DB."HIGH LEVEL VALUE (H)" AT %DB2223.DBD30, 1 s
   "PIT424_RIO6_ALM_ANALOG_DB_LOW LEVEL VALUE (L)" : Real = PLC PIT424_RIO6_ALM_ANALOG_DB."LOW LEVEL VALUE (L)" AT %DB2223.DBD26, 1 s
   "PIT424_RIO6_ALM_ANALOG_DB_VERY HIGH LEVEL VALUE (HH)" : Real = PLC PIT424_RIO6_ALM_ANALOG_DB."VERY HIGH LEVEL VALUE (HH)" AT %DB2223.DBD34, 1 s
   "PIT424_RIO6_ALM_ANALOG_DB_VERY LOW LEVEL VALUE (LL)" : Real = PLC PIT424_RIO6_ALM_ANALOG_DB."VERY LOW LEVEL VALUE (LL)" AT %DB2223.DBD22, 1 s
   "PIT424_RIO7_ALM_ANALOG_DB_HIGH LEVEL VALUE (H)" : Real = PLC PIT424_RIO7_ALM_ANALOG_DB."HIGH LEVEL VALUE (H)" AT %DB2224.DBD30, 1 s
   "PIT424_RIO7_ALM_ANALOG_DB_LOW LEVEL VALUE (L)" : Real = PLC PIT424_RIO7_ALM_ANALOG_DB."LOW LEVEL VALUE (L)" AT %DB2224.DBD26, 1 s
   "PIT424_RIO7_ALM_ANALOG_DB_VERY HIGH LEVEL VALUE (HH)" : Real = PLC PIT424_RIO7_ALM_ANALOG_DB."VERY HIGH LEVEL VALUE (HH)" AT %DB2224.DBD34, 1 s
   "PIT424_RIO7_ALM_ANALOG_DB_VERY LOW LEVEL VALUE (LL)" : Real = PLC PIT424_RIO7_ALM_ANALOG_DB."VERY LOW LEVEL VALUE (LL)" AT %DB2224.DBD22, 1 s
   "PIT424PORT_ALM_ANALOG_DB_HIGH LEVEL VALUE (H)" : Real = PLC PIT424PORT_ALM_ANALOG_DB."HIGH LEVEL VALUE (H)" AT %DB2070.DBD30, 1 s
   "PIT424PORT_ALM_ANALOG_DB_LOW LEVEL VALUE (L)" : Real = PLC PIT424PORT_ALM_ANALOG_DB."LOW LEVEL VALUE (L)" AT %DB2070.DBD26, 1 s
   "PIT424PORT_ALM_ANALOG_DB_VERY HIGH LEVEL VALUE (HH)" : Real = PLC PIT424PORT_ALM_ANALOG_DB."VERY HIGH LEVEL VALUE (HH)" AT %DB2070.DBD34, 1 s
   "PIT424PORT_ALM_ANALOG_DB_VERY LOW LEVEL VALUE (LL)" : Real = PLC PIT424PORT_ALM_ANALOG_DB."VERY LOW LEVEL VALUE (LL)" AT %DB2070.DBD22, 1 s
   "Pre Dwell Time Remains" : Int = PLC "2102_TIME_CALCS_DB"."PRE-DWEL HOURS REMNG" AT %DB1.DBW0, 1 s
   "Process Gas Compressor Running/Stopped" : Bool = PLC "Process Gas Compressor Running/Stopped" AT %I139.0, 1 s
   "PT415_FPT_ALM_ANALOG_DB_HIGH LEVEL VALUE (H)" : Real = PLC PT415_FPT_ALM_ANALOG_DB."HIGH LEVEL VALUE (H)" AT %DB2213.DBD30, 1 s
   "PT415_FPT_ALM_ANALOG_DB_LOW LEVEL VALUE (L)" : Real = PLC PT415_FPT_ALM_ANALOG_DB."LOW LEVEL VALUE (L)" AT %DB2213.DBD26, 1 s
   "PT415_FPT_ALM_ANALOG_DB_VERY HIGH LEVEL VALUE (HH)" : Real = PLC PT415_FPT_ALM_ANALOG_DB."VERY HIGH LEVEL VALUE (HH)" AT %DB2213.DBD34, 1 s
   "PT415_FPT_ALM_ANALOG_DB_VERY LOW LEVEL VALUE (LL)" : Real = PLC PT415_FPT_ALM_ANALOG_DB."VERY LOW LEVEL VALUE (LL)" AT %DB2213.DBD22, 1 s
   "PT415_RIO3_ALM_ANALOG_DB_HIGH LEVEL VALUE (H)" : Real = PLC PT415_RIO3_ALM_ANALOG_DB."HIGH LEVEL VALUE (H)" AT %DB2215.DBD30, 1 s
   "PT415_RIO3_ALM_ANALOG_DB_LOW LEVEL VALUE (L)" : Real = PLC PT415_RIO3_ALM_ANALOG_DB."LOW LEVEL VALUE (L)" AT %DB2215.DBD26, 1 s
   "PT415_RIO3_ALM_ANALOG_DB_VERY HIGH LEVEL VALUE (HH)" : Real = PLC PT415_RIO3_ALM_ANALOG_DB."VERY HIGH LEVEL VALUE (HH)" AT %DB2215.DBD34, 1 s
   "PT415_RIO3_ALM_ANALOG_DB_VERY LOW LEVEL VALUE (LL)" : Real = PLC PT415_RIO3_ALM_ANALOG_DB."VERY LOW LEVEL VALUE (LL)" AT %DB2215.DBD22, 1 s
   "PT415_RIO4_ALM_ANALOG_DB_HIGH LEVEL VALUE (H)" : Real = PLC PT415_RIO4_ALM_ANALOG_DB."HIGH LEVEL VALUE (H)" AT %DB2216.DBD30, 1 s
   "PT415_RIO4_ALM_ANALOG_DB_LOW LEVEL VALUE (L)" : Real = PLC PT415_RIO4_ALM_ANALOG_DB."LOW LEVEL VALUE (L)" AT %DB2216.DBD26, 1 s
   "PT415_RIO4_ALM_ANALOG_DB_VERY HIGH LEVEL VALUE (HH)" : Real = PLC PT415_RIO4_ALM_ANALOG_DB."VERY HIGH LEVEL VALUE (HH)" AT %DB2216.DBD34, 1 s
   "PT415_RIO4_ALM_ANALOG_DB_VERY LOW LEVEL VALUE (LL)" : Real = PLC PT415_RIO4_ALM_ANALOG_DB."VERY LOW LEVEL VALUE (LL)" AT %DB2216.DBD22, 1 s
   "PT415_RIO5_ALM_ANALOG_DB_HIGH LEVEL VALUE (H)" : Real = PLC PT415_RIO5_ALM_ANALOG_DB."HIGH LEVEL VALUE (H)" AT %DB2217.DBD30, 1 s
   "PT415_RIO5_ALM_ANALOG_DB_LOW LEVEL VALUE (L)" : Real = PLC PT415_RIO5_ALM_ANALOG_DB."LOW LEVEL VALUE (L)" AT %DB2217.DBD26, 1 s
   "PT415_RIO5_ALM_ANALOG_DB_VERY HIGH LEVEL VALUE (HH)" : Real = PLC PT415_RIO5_ALM_ANALOG_DB."VERY HIGH LEVEL VALUE (HH)" AT %DB2217.DBD34, 1 s
   "PT415_RIO5_ALM_ANALOG_DB_VERY LOW LEVEL VALUE (LL)" : Real = PLC PT415_RIO5_ALM_ANALOG_DB."VERY LOW LEVEL VALUE (LL)" AT %DB2217.DBD22, 1 s
   "PT415_RIO6_ALM_ANALOG_DB_HIGH LEVEL VALUE (H)" : Real = PLC PT415_RIO6_ALM_ANALOG_DB."HIGH LEVEL VALUE (H)" AT %DB2218.DBD30, 1 s
   "PT415_RIO6_ALM_ANALOG_DB_LOW LEVEL VALUE (L)" : Real = PLC PT415_RIO6_ALM_ANALOG_DB."LOW LEVEL VALUE (L)" AT %DB2218.DBD26, 1 s
   "PT415_RIO6_ALM_ANALOG_DB_VERY HIGH LEVEL VALUE (HH)" : Real = PLC PT415_RIO6_ALM_ANALOG_DB."VERY HIGH LEVEL VALUE (HH)" AT %DB2218.DBD34, 1 s
   "PT415_RIO6_ALM_ANALOG_DB_VERY LOW LEVEL VALUE (LL)" : Real = PLC PT415_RIO6_ALM_ANALOG_DB."VERY LOW LEVEL VALUE (LL)" AT %DB2218.DBD22, 1 s
   "PT415_RIO7_ALM_ANALOG_DB_HIGH LEVEL VALUE (H)" : Real = PLC PT415_RIO7_ALM_ANALOG_DB."HIGH LEVEL VALUE (H)" AT %DB2225.DBD30, 1 s
   "PT415_RIO7_ALM_ANALOG_DB_LOW LEVEL VALUE (L)" : Real = PLC PT415_RIO7_ALM_ANALOG_DB."LOW LEVEL VALUE (L)" AT %DB2225.DBD26, 1 s
   "PT415_RIO7_ALM_ANALOG_DB_VERY HIGH LEVEL VALUE (HH)" : Real = PLC PT415_RIO7_ALM_ANALOG_DB."VERY HIGH LEVEL VALUE (HH)" AT %DB2225.DBD34, 1 s
   "PT415_RIO7_ALM_ANALOG_DB_VERY LOW LEVEL VALUE (LL)" : Real = PLC PT415_RIO7_ALM_ANALOG_DB."VERY LOW LEVEL VALUE (LL)" AT %DB2225.DBD22, 1 s
   "PT415PORT_ALM_ANALOG_DB_HIGH LEVEL VALUE (H)" : Real = PLC PT415PORT_ALM_ANALOG_DB."HIGH LEVEL VALUE (H)" AT %DB2069.DBD30, 1 s
   "PT415PORT_ALM_ANALOG_DB_LOW LEVEL VALUE (L)" : Real = PLC PT415PORT_ALM_ANALOG_DB."LOW LEVEL VALUE (L)" AT %DB2069.DBD26, 1 s
   "PT415PORT_ALM_ANALOG_DB_VERY HIGH LEVEL VALUE (HH)" : Real = PLC PT415PORT_ALM_ANALOG_DB."VERY HIGH LEVEL VALUE (HH)" AT %DB2069.DBD34, 1 s
   "PT415PORT_ALM_ANALOG_DB_VERY LOW LEVEL VALUE (LL)" : Real = PLC PT415PORT_ALM_ANALOG_DB."VERY LOW LEVEL VALUE (LL)" AT %DB2069.DBD22, 1 s
   "R1_SPR_AI_126" : Real = PLC "12_AI_Data".R1_SPR_AI_126_SCALED AT %DB1.DBX0.0, 1 s
   "R1_SPR_AI_132" : Real = PLC "12_AI_Data".R1_SPR_AI_132_SCALED AT %DB1.DBD0, 1 s
   "R1_SPR_AQ_102" : Real = PLC "16_AQ_Data".R1_SPR_AQ_102 AT %DB1.DBD0, 1 s
   "R1_SPR_AQ_104" : Real = PLC "16_AQ_Data".R1_SPR_AQ_104 AT %DB1.DBD0, 1 s
   "R1_SPR_DI_3_7" : Bool = PLC "10_DI_Data".R1_SPR_DI_3_7 AT %DB1.DBX0.0, 1 s
   "R2_SPR_AQ_96" : Real = PLC "16_AQ_Data".R2_SPR_AQ_96 AT %DB1.DBD0, 1 s
   "R2_SPR_AQ_98" : Real = PLC "16_AQ_Data".R2_SPR_AQ_98 AT %DB1.DBD0, 1 s
   "R2_SPR_DI_0_2" : Bool = PLC "10 DI_DATA".R2_SPR_DI_0_2 AT %DB1.DBX0.0, 1 s
   "R2_SPR_DI_0_3" : Bool = PLC "10 DI_DATA".R2_SPR_DI_0_3 AT %DB1.DBX0.0, 1 s
   "R2_SPR_DI_1_6 Spare Input" : Bool = PLC "10 DI_DATA".R2_SPR_DI_1_6 AT %DB1.DBX0.0, 1 s
   "R2_SPR_DI_3_2" : Bool = PLC "10 DI_DATA".R2_SPR_DI_3_2 AT %DB1.DBX0.0, 1 s
   "R2_SPR_DI_3_7" : Bool = PLC "10 DI_DATA".R2_SPR_DI_3_7 AT %DB1.DBX0.0, 1 s
   "RESET_STEP" : Bool = PLC RESET_STEP AT %M12.0, 1 s
   "RIO1 Tanks Pressure Switch Hi Hi" : Bool = PLC "RIO1 Tanks Pressure Switch Hi Hi" AT %I9.1, 1 s
   "RIO1_SPR_DI_0_6" : Bool = PLC RIO1_SPR_DI_0_6 AT %I0.6, 1 s
   "RIO1_SPR_DI_0_7" : Bool = PLC RIO1_SPR_DI_0_7 AT %I0.7, 1 s
   "RIO1_SPR_DI_3_6" : Bool = PLC RIO1_SPR_DI_3_6 AT %I3.6, 1 s
   "RIO1_SPR_DI_3_7" : Bool = PLC RIO1_SPR_DI_3_7 AT %I3.7, 1 s
   "RIO1_SPR_DI_6_6" : Bool = PLC RIO1_SPR_DI_6_6 AT %I6.6, 1 s
   "RIO1_SPR_DI_6_7" : Bool = PLC RIO1_SPR_DI_6_7 AT %I6.7, 1 s
   "RIO1_SPR_DI_9_4" : Bool = PLC RIO1_SPR_DI_9_4 AT %I9.4, 1 s
   "RIO1_SPR_DI_9_5" : Bool = PLC RIO1_SPR_DI_9_5 AT %I9.5, 1 s
   "RIO1_SPR_DI_9_6" : Bool = PLC RIO1_SPR_DI_9_6 AT %I9.6, 1 s
   "RIO1_SPR_DI_9_7" : Bool = PLC RIO1_SPR_DI_9_7 AT %I9.7, 1 s
   "RIO2 Tanks Pressure Switch Hi Hi" : Bool = PLC "RIO2 Tanks Pressure Switch Hi Hi" AT %I21.1, 1 s
   "RIO2_SPR_DI_15_6" : Bool = PLC RIO2_SPR_DI_15_6 AT %I15.6, 1 s
   "RIO2_SPR_DI_15_7" : Bool = PLC RIO2_SPR_DI_15_7 AT %I15.7, 1 s
   "RIO2_SPR_DI_18_6" : Bool = PLC RIO2_SPR_DI_18_6 AT %I18.6, 1 s
   "RIO2_SPR_DI_18_7" : Bool = PLC RIO2_SPR_DI_18_7 AT %I18.7, 1 s
   "RIO2_SPR_DI_21_3" : Bool = PLC RIO2_SPR_DI_21_3 AT %I21.3, 1 s
   "RIO2_SPR_DI_21_4" : Bool = PLC RIO2_SPR_DI_21_4 AT %I21.4, 1 s
   "RIO2_SPR_DI_21_5" : Bool = PLC RIO2_SPR_DI_21_5 AT %I21.5, 1 s
   "RIO2_SPR_DI_21_6" : Bool = PLC RIO2_SPR_DI_21_6 AT %I21.6, 1 s
   "RIO2_SPR_DI_21_7" : Bool = PLC RIO2_SPR_DI_21_7 AT %I21.7, 1 s